// TIA Portal project "e009004v439" (V15.1) (continued)
HMI tags "Tag table_7"
   "Receta Almacén 2\Recetas.REC_MG2.C" : DInt AT %DB51.DBD182, 1 s   // Mot Piece : Côte C
   "Receta Almacén 2\CA_KM01_2" : Bool AT %M19.4, 1 s   // Intercambiador Almacenes Retroceso (Alm2)
   "Receta Almacén 2\OFFSET.REC_MG2.OFFSET_F4" : Int AT %DB52.DBW66, 1 s   // Punto de Formado 4
   "Receta Almacén 2\DB_OP.M2_XCPT" : Bool AT %DB50.DBX382.0, 1 s   // Almacén 2 Entrega Pieza
   "Receta Almacén 2\Detalles" : Bool, internal
   "Receta Almacén 2\DB_OP.M2.MPP" : Bool AT %DB50.DBX420.0, 1 s   // Presencia de Pieza
   "Receta Almacén 2\OFFSET.REC_MG2.OFFSET_F1" : Int AT %DB52.DBW60, 1 s   // Punto de Formado 1
   "Receta Almacén 2\Recetas.REC_MG2.A" : DInt AT %DB51.DBD174, 1 s   // Mot Piece : Côte A
   "Receta Almacén 2\OFFSET.REC_MG2.OFFSET_PL2_1" : Int AT %DB52.DBW72, 1 s   // Plegador 2 Pliego 1
   "Receta Almacén 2\Recetas.REC_MG2.NOM" : String[8] AT %DB51.DBX160.0, 1 s
   "Receta Almacén 2\Recetas.REC_MG2.B" : DInt AT %DB51.DBD178, 1 s   // Mot Piece : Côte B
   "Receta Almacén 2\VerHeladera" : Bool, internal
   "Receta Almacén 2\OFFSET.REC_MG2.OFFSET_F2" : Int AT %DB52.DBW62, 1 s   // Punto de Formado 2
   "Receta Almacén 2\Recetas.REC_MG2.D" : DInt AT %DB51.DBD186, 1 s   // Mot Piece : Côte D
   "Receta Almacén 2\OFFSET.REC_MG2.OFFSET_PL2_2" : Int AT %DB52.DBW74, 1 s   // Plegador 2 Pliego 2
   "Receta Almacén 2\26S6" : Bool AT %I3.5, 1 s   // Presencia de Almacén 2 en Puesto de Espera
   "Receta Almacén 2\OFFSET.REC_MG2.OFFSET_PL1_1" : Int AT %DB52.DBW68, 1 s   // Plegador 1 Pliego 1
   "Receta Almacén 2\OFFSET.REC_MG2.OFFSET_F3" : Int AT %DB52.DBW64, 1 s   // Punto de Formado 3
   "Receta Almacén 2\OFFSET.REC_MG2.OFFSET_PL1_2" : Int AT %DB52.DBW70, 1 s   // Plegador 1 Pliego 2

HMI tags "PiezaPerfiladores"
   "Perfiladores\Perfilador.B" : Int AT %DB8.DBW2, 1 s
   "Perfiladores\Perfilador.PresenciaPieza" : Bool AT %DB8.DBX46.0, 1 s
   "Perfiladores\Perfilador.F1" : Int AT %DB8.DBW8, 1 s
   "Perfiladores\Perfilador.F3" : Int AT %DB8.DBW12, 1 s
   "Perfiladores\Perfilador.PL2_1" : Int AT %DB8.DBW20, 1 s
   "Perfiladores\Perfilador.PL1_1" : Int AT %DB8.DBW16, 1 s
   "Perfiladores\Perfilador.C" : Int AT %DB8.DBW4, 1 s
   "Perfiladores\Perfilador.PL1_2" : Int AT %DB8.DBW18, 1 s
   "Perfiladores\Perfilador.F2" : Int AT %DB8.DBW10, 1 s
   "Perfiladores\Perfilador.F4" : Int AT %DB8.DBW14, 1 s
   "Perfiladores\Perfilador.A" : Int AT %DB8.DBW0, 1 s
   "Perfiladores\Perfilador.PL2_2" : Int AT %DB8.DBW22, 1 s
   "Perfiladores\Perfilador.D" : Int AT %DB8.DBW6, 1 s
   "Forz_Transf-3" : Bool AT %M113.2, 1 s
   "Forz_Transf2" : Bool AT %M113.1, 1 s
   "Forz_Transf1" : Bool AT %M113.0, 1 s
   "Perfiladores\Perfilador.Nombre" : String[20] AT %DB8.DBX24.0, 1 s

HMI tags "PiezaCinta"
   "Cinta\Cinta.PresenciaPieza" : Bool AT %DB9.DBX46.0, 1 s
   "Cinta\Cinta.PL2_1" : Int AT %DB9.DBW20, 1 s
   "Cinta\Cinta.C" : Int AT %DB9.DBW4, 1 s
   "Cinta\Cinta.A" : Int AT %DB9.DBW0, 1 s
   "Cinta\Cinta.F4" : Int AT %DB9.DBW14, 1 s
   "Cinta\Cinta.F3" : Int AT %DB9.DBW12, 1 s
   "Cinta\Cinta.PL2_2" : Int AT %DB9.DBW22, 1 s
   "Cinta\Cinta.PL1_1" : Int AT %DB9.DBW16, 1 s
   "Cinta\Cinta.PL1_2" : Int AT %DB9.DBW18, 1 s
   "Cinta\Cinta.F2" : Int AT %DB9.DBW10, 1 s
   "Cinta\Cinta.D" : Int AT %DB9.DBW6, 1 s
   "Cinta\Cinta.B" : Int AT %DB9.DBW2, 1 s
   "Cinta\Cinta.F1" : Int AT %DB9.DBW8, 1 s
   "Cinta\Cinta.Nombre" : String[20] AT %DB9.DBX24.0, 1 s

HMI tags "PiezaAlm2"
   "Almacén 2\PAlmacén.F3" : Int AT %DB5.DBW12, 1 s
   "Almacén 2\PAlmacén.B" : Int AT %DB5.DBW2, 1 s
   "Almacén 2\PAlmacén.PL2_1" : Int AT %DB5.DBW20, 1 s
   "Almacén 2\PAlmacén.PresenciaPieza" : Bool AT %DB5.DBX46.0, 1 s
   "Almacén 2\PAlmacén.F1" : Int AT %DB5.DBW8, 1 s
   "Almacén 2\PAlmacén.PL2_2" : Int AT %DB5.DBW22, 1 s
   "Almacén 2\PAlmacén.A" : Int AT %DB5.DBW0, 1 s
   "Almacén 2\PAlmacén.F2" : Int AT %DB5.DBW10, 1 s
   "Almacén 2\PAlmacén.F4" : Int AT %DB5.DBW14, 1 s
   "Almacén 2\PAlmacén.C" : Int AT %DB5.DBW4, 1 s
   "Almacén 2\PAlmacén.PL1_1" : Int AT %DB5.DBW16, 1 s
   "Almacén 2\PAlmacén.PL1_2" : Int AT %DB5.DBW18, 1 s
   "Almacén 2\PAlmacén.D" : Int AT %DB5.DBW6, 1 s
   "Almacén 2\PAlmacén.Nombre" : String[20] AT %DB5.DBX24.0, 1 s

HMI tags "PiezaAlm1"
   "Almacén 1\PAlmacén.PL2_2" : Int AT %DB4.DBW22, 1 s
   "Almacén 1\PAlmacén.PL2_1" : Int AT %DB4.DBW20, 1 s
   "Almacén 1\PAlmacén.D" : Int AT %DB4.DBW6, 1 s
   "Almacén 1\PAlmacén.A" : Int AT %DB4.DBW0, 1 s
   "Almacén 1\PAlmacén.F4" : Int AT %DB4.DBW14, 1 s
   "Almacén 1\PAlmacén.B" : Int AT %DB4.DBW2, 1 s
   "Almacén 1\PAlmacén.F3" : Int AT %DB4.DBW12, 1 s
   "Almacén 1\PAlmacén.F2" : Int AT %DB4.DBW10, 1 s
   "Almacén 1\PAlmacén.PL1_2" : Int AT %DB4.DBW18, 1 s
   "Almacén 1\PAlmacén.F1" : Int AT %DB4.DBW8, 1 s
   "Almacén 1\PAlmacén.C" : Int AT %DB4.DBW4, 1 s
   "Almacén 1\PAlmacén.PL1_1" : Int AT %DB4.DBW16, 1 s
   "Almacén 1\PAlmacén.Nombre" : String[20] AT %DB4.DBX24.0, 1 s
   "PL_Resoluc_INCDECF" : Int AT %DB19.DBW8, 1 s
   "PL_Resoluc_INCDECPL" : Int AT %DB19.DBW18, 1 s
   "Almacén 1\PAlmacén.PresenciaPieza_1" : Bool AT %DB4.DBX46.1, 1 s

HMI tags "Alarmas"
   "Alarma 1" : Bool AT %DB50.DBX80.0, 1 s
   "Alarma 2" : Bool AT %DB50.DBX80.1, 1 s
   "Alarma 3" : Bool AT %DB50.DBX80.2, 1 s
   "Alarma 4" : Bool AT %DB50.DBX80.3, 1 s
   "Alarma 5" : Bool AT %DB50.DBX80.4, 1 s
   "Alarma 6" : Bool AT %DB50.DBX80.5, 1 s
   "Alarma 7" : Bool AT %DB50.DBX80.6, 1 s
   "Alarma 8" : Bool AT %DB50.DBX80.7, 1 s
   "Alarma 9" : Bool AT %DB50.DBX81.0, 1 s
   "Alarma 10" : Bool AT %DB50.DBX81.1, 1 s
   "Alarma 11" : Bool AT %DB50.DBX81.2, 1 s
   "Alarma 12" : Bool AT %DB50.DBX81.3, 1 s
   "Alarma 13" : Bool AT %DB50.DBX81.4, 1 s
   "Alarma 14" : Bool AT %DB50.DBX81.5, 1 s
   "Alarma 15" : Bool AT %DB50.DBX81.6, 1 s
   "Alarma 16" : Bool AT %DB50.DBX81.7, 1 s
   "Alarma 17" : Bool AT %DB50.DBX82.0, 1 s
   "Alarma 18" : Bool AT %DB50.DBX82.1, 1 s
   "Alarma 19" : Bool AT %DB50.DBX82.2, 1 s
   "Alarma 20" : Bool AT %DB50.DBX82.3, 1 s
   "Alarma 21" : Bool AT %DB50.DBX82.4, 1 s
   "Alarma 22" : Bool AT %DB50.DBX82.5, 1 s
   "Alarma 23" : Bool AT %DB50.DBX82.6, 1 s
   "Alarma 24" : Bool AT %DB50.DBX82.7, 1 s
   "Alarma 25" : Bool AT %DB50.DBX83.0, 1 s
   "Alarma 26" : Bool AT %DB50.DBX83.1, 1 s
   "Alarma 27" : Bool AT %DB50.DBX83.2, 1 s
   "Alarma 28" : Bool AT %DB50.DBX83.3, 1 s
   "Alarma 29" : Bool AT %DB50.DBX83.4, 1 s
   "Alarma 30" : Bool AT %DB50.DBX83.5, 1 s
   "Alarma 31" : Bool AT %DB50.DBX83.6, 1 s
   "Alarma 32" : Bool AT %DB50.DBX83.7, 1 s
   "Alarma 33" : Bool AT %DB50.DBX84.0, 1 s
   "Alarma 34" : Bool AT %DB50.DBX84.1, 1 s
   "Alarma 35" : Bool AT %DB50.DBX84.2, 1 s
   "Alarma 36" : Bool AT %DB50.DBX84.3, 1 s
   "Alarma 37" : Bool AT %DB50.DBX84.4, 1 s
   "Alarma 38" : Bool AT %DB50.DBX84.5, 1 s
   "Alarma 39" : Bool AT %DB50.DBX84.6, 1 s
   "Alarma 40" : Bool AT %DB50.DBX84.7, 1 s
   "Alarma 41" : Bool AT %DB50.DBX85.0, 1 s
   "Alarma 42" : Bool AT %DB50.DBX85.1, 1 s
   "Alarma 43" : Bool AT %DB50.DBX85.2, 1 s
   "Alarma 44" : Bool AT %DB50.DBX85.3, 1 s
   "Alarma 45" : Bool AT %DB50.DBX85.4, 1 s
   "Alarma 46" : Bool AT %DB50.DBX85.5, 1 s
   "Alarma 47" : Bool AT %DB50.DBX85.6, 1 s
   "Alarma 48" : Bool AT %DB50.DBX85.7, 1 s
   "Alarma 49" : Bool AT %DB50.DBX86.0, 1 s
   "Alarma 50" : Bool AT %DB50.DBX86.1, 1 s
   "Alarma 51" : Bool AT %DB50.DBX86.2, 1 s
   "Alarma 52" : Bool AT %DB50.DBX86.3, 1 s
   "Alarma 53" : Bool AT %DB50.DBX86.4, 1 s
   "Alarma 54" : Bool AT %DB50.DBX86.5, 1 s
   "Alarma 55" : Bool AT %DB50.DBX86.6, 1 s
   "Alarma 56" : Bool AT %DB50.DBX86.7, 1 s
   "Alarma 57" : Bool AT %DB50.DBX87.0, 1 s
   "Alarma 58" : Bool AT %DB50.DBX87.1, 1 s
   "Alarma 59" : Bool AT %DB50.DBX87.2, 1 s
   "Alarma 60" : Bool AT %DB50.DBX87.3, 1 s
   "Alarma 61" : Bool AT %DB50.DBX87.4, 1 s
   "Alarma 62" : Bool AT %DB50.DBX87.5, 1 s
   "Alarma 63" : Bool AT %DB50.DBX87.6, 1 s
   "Alarma 64" : Bool AT %DB50.DBX87.7, 1 s
   "Alarma 65" : Bool AT %DB50.DBX88.0, 1 s
   "Alarma 66" : Bool AT %DB50.DBX88.1, 1 s
   "Alarma 67" : Bool AT %DB50.DBX88.2, 1 s
   "Alarma 68" : Bool AT %DB50.DBX88.3, 1 s
   "Alarma 69" : Bool AT %DB50.DBX88.4, 1 s
   "Alarma 70" : Bool AT %DB50.DBX88.5, 1 s
   "Alarma 71" : Bool AT %DB50.DBX88.6, 1 s
   "Alarma 72" : Bool AT %DB50.DBX88.7, 1 s
   "Alarma 73" : Bool AT %DB50.DBX89.0, 1 s
   "Alarma 74" : Bool AT %DB50.DBX89.1, 1 s
   "Alarma 75" : Bool AT %DB50.DBX89.2, 1 s
   "Alarma 76" : Bool AT %DB50.DBX89.3, 1 s
   "Alarma 77" : Bool AT %DB50.DBX89.4, 1 s
   "Alarma 78" : Bool AT %DB50.DBX89.5, 1 s
   "Alarma 79" : Bool AT %DB50.DBX89.6, 1 s
   "Alarma 80" : Bool AT %DB50.DBX89.7, 1 s
   "Alarma 81" : Bool AT %DB50.DBX90.0, 1 s
   "Alarma 82" : Bool AT %DB50.DBX90.1, 1 s
   "Alarma 83" : Bool AT %DB50.DBX90.2, 1 s
   "Alarma 84" : Bool AT %DB50.DBX90.3, 1 s
   "Alarma 85" : Bool AT %DB50.DBX90.4, 1 s
   "Alarma 86" : Bool AT %DB50.DBX90.5, 1 s
   "Alarma 87" : Bool AT %DB50.DBX90.6, 1 s
   "Alarma 88" : Bool AT %DB50.DBX90.7, 1 s
   "Alarma 89" : Bool AT %DB50.DBX91.0, 1 s
   "Alarma 90" : Bool AT %DB50.DBX91.1, 1 s
   "Alarma 91" : Bool AT %DB50.DBX91.2, 1 s
   "Alarma 92" : Bool AT %DB50.DBX91.3, 1 s
   "Alarma 93" : Bool AT %DB50.DBX91.4, 1 s
   "Alarma 94" : Bool AT %DB50.DBX91.5, 1 s
   "Alarma 95" : Bool AT %DB50.DBX91.6, 1 s
   "Alarma 96" : Bool AT %DB50.DBX91.7, 1 s
   "Alarma 97" : Bool AT %DB50.DBX92.0, 1 s
   "Alarma 98" : Bool AT %DB50.DBX92.1, 1 s
   "Alarma 99" : Bool AT %DB50.DBX92.2, 1 s
   "Alarma 100" : Bool AT %DB50.DBX92.3, 1 s
   "Alarma 101" : Bool AT %DB50.DBX92.4, 1 s
   "Alarma 102" : Bool AT %DB50.DBX92.5, 1 s
   "Alarma 103" : Bool AT %DB50.DBX92.6, 1 s
   "Alarma 104" : Bool AT %DB50.DBX92.7, 1 s
   "Alarma 105" : Bool AT %DB50.DBX93.0, 1 s
   "Alarma 106" : Bool AT %DB50.DBX93.1, 1 s
   "Alarma 107" : Bool AT %DB50.DBX93.2, 1 s
   "Alarma 108" : Bool AT %DB50.DBX93.3, 1 s
   "Alarma 109" : Bool AT %DB50.DBX93.4, 1 s
   "Alarma 110" : Bool AT %DB50.DBX93.5, 1 s
   "Alarma 111" : Bool AT %DB50.DBX93.6, 1 s
   "Alarma 112" : Bool AT %DB50.DBX93.7, 1 s
   "Alarma 113" : Bool AT %DB50.DBX94.0, 1 s
   "Alarma 114" : Bool AT %DB50.DBX94.1, 1 s
   "Alarma 115" : Bool AT %DB50.DBX94.2, 1 s
   "Alarma 116" : Bool AT %DB50.DBX94.3, 1 s
   "Alarma 117" : Bool AT %DB50.DBX94.4, 1 s
   "Alarma 118" : Bool AT %DB50.DBX94.5, 1 s
   "Alarma 119" : Bool AT %DB50.DBX94.6, 1 s
   "Alarma 120" : Bool AT %DB50.DBX94.7, 1 s
   "Alarma 121" : Bool AT %DB50.DBX95.0, 1 s
   "PL1_Pos00" : Bool AT %DB50.DBX393.0, 1 s

HMI tags "Atasco Perfilador"
   "Sensor 1" : Bool AT %I14.4, 100 ms
   "Sensor 2" : Bool AT %I14.5, 100 ms
   "Sensor 3" : Bool AT %I14.6, 100 ms
   "Sensor 4" : Bool AT %I14.7, 100 ms
   "Sensor 5" : Bool AT %I18.3, 100 ms
   "Sensor 6" : Bool AT %I16.0, 100 ms
   "Sensor 7" : Bool AT %I16.1, 100 ms
   "Sensor 8" : Bool AT %I16.2, 100 ms
   "Sensor 9" : Bool AT %I16.3, 100 ms
   "Sensor 10" : Bool AT %I16.4, 100 ms
   "Sensor 11" : Bool AT %I16.5, 100 ms
   "Sensor 12" : Bool AT %I16.6, 100 ms
   "Sensor 13" : Bool AT %I16.7, 100 ms
   "Sensor 14" : Bool AT %I17.0, 100 ms
   "Sensor 15" : Bool AT %I17.1, 100 ms
   "Sensor 16" : Bool AT %I17.2, 100 ms
   "Sensor 17" : Bool AT %I17.3, 100 ms
   "Sensor 18" : Bool AT %I17.4, 100 ms
   "Sensor 19" : Bool AT %I17.5, 100 ms
   "Sensor 20" : Bool, internal
   "Sensor 21" : Bool AT %I17.6, 100 ms
   "Sensor 22" : Bool AT %I18.0, 100 ms
   "Sensor 23" : Bool AT %I18.1, 100 ms
   "Sensor 24" : Bool AT %I18.2, 100 ms
   "36S10" : Bool AT %I15.0, 1 s

HMI tags "PiezaDescargador"
   "Descargador-A" : Int AT %DB12.DBW0, 1 s
   "Descargador-B" : Int AT %DB12.DBW2, 1 s
   "Descargador-C" : Int AT %DB12.DBW4, 1 s
   "Descargador-D" : Int AT %DB12.DBW6, 1 s
   "Descargador-F1" : Int AT %DB12.DBW8, 1 s
   "Descargador-F2" : Int AT %DB12.DBW10, 1 s
   "Descargador-F3" : Int AT %DB12.DBW12, 1 s
   "Descargador-F4" : Int AT %DB12.DBW14, 1 s
   "Descargador-PL1_1" : Int AT %DB12.DBW16, 1 s
   "Descargador-PL1_2" : Int AT %DB12.DBW18, 1 s
   "Descargador-PL2_1" : Int AT %DB12.DBW20, 1 s
   "Descargador-PL2_2" : Int AT %DB12.DBW22, 1 s
   "Descargador-Nombre" : String[20] AT %DB12.DBX24.0, 1 s
   "Descargador-PiezaPresente" : Bool AT %DB12.DBX46.0, 1 s
   "Descargador-Almacen" : Bool AT %DB12.DBX46.1, 1 s
   "Descargador-PL2_3" : Int AT %DB12.DBW24, 1 s

HMI tags "ProcesoPlegadores"
   "PL_Estados" : Int AT %MW150, 1 s
   "PL_Concatenadoras" : Int AT %MW152, 1 s
   "PL_S_0" : Bool AT %M150.0, 1 s
   "PL_S_1" : Bool AT %M150.1, 1 s
   "PL_S_2" : Bool AT %M150.2, 1 s
   "PL_S_3" : Bool AT %M150.3, 1 s
   "PL_S_4" : Bool AT %M150.4, 1 s
   "PL_S_5" : Bool AT %M150.5, 1 s
   "PL_S_6" : Bool AT %M150.6, 1 s
   "PL_S_7" : Bool AT %M150.7, 1 s
   "PL_S_8" : Bool AT %M151.0, 1 s
   "PL_S_9" : Bool AT %M151.1, 1 s
   "PL_S_10" : Bool AT %M151.2, 1 s
   "PL_S_11" : Bool AT %M151.3, 1 s
   "PL_S_12" : Bool AT %M151.4, 1 s
   "PL_S_13" : Bool AT %M151.5, 1 s
   "PL_S_14" : Bool AT %M151.6, 1 s
   "PL_S_15" : Bool AT %M151.7, 1 s
   "STOP_RUN" : Bool AT %M101.3, 1 s
   "PL_Continuar" : Bool AT %M101.4, 1 s
   "PL_Reset" : Bool AT %M101.5, 1 s
   "PL_en_Ciclo" : Bool AT %M10.3, 1 s
   "PL_Prioritarias" : Int AT %MW154, 1 s
   "PL_P_0" : Bool AT %M154.0, 1 s
   "PL_P_1" : Bool AT %M154.1, 1 s
   "PL_P_2" : Bool AT %M154.2, 1 s
   "PL_P_3" : Bool AT %M154.3, 1 s
   "PL_P_4" : Bool AT %M154.4, 1 s
   "PL_P_5" : Bool AT %M154.5, 1 s
   "PL_P_6" : Bool AT %M154.6, 1 s
   "PL_P_7" : Bool AT %M154.7, 1 s
   "PL_P_8" : Bool AT %M155.0, 1 s
   "PL_P_9" : Bool AT %M155.1, 1 s
   "PL_P_10" : Bool AT %M155.2, 1 s
   "PL_P_11" : Bool AT %M155.3, 1 s
   "PL_P_12" : Bool AT %M155.4, 1 s
   "PL_P_13" : Bool AT %M155.5, 1 s
   "PL_P_14" : Bool AT %M155.6, 1 s
   "PL_P_15" : Bool AT %M155.7, 1 s
   "PL_Req_Pos_Recep" : Bool AT %M100.0, 1 s
   "PL_Req_Pos_Pleg1" : Bool AT %M100.1, 1 s
   "PL_Req_Pos_Pleg2" : Bool AT %M100.3, 1 s
   "PL_Req_Pos_Entrega" : Bool AT %M100.4, 1 s
   "PL_Req_Pos_Espera" : Bool AT %M100.5, 1 s
   "PL_En_Pos_Espera" : Bool AT %M180.0, 1 s
   "PL_En_Pos_Recepción" : Bool AT %M180.1, 1 s
   "PL_En_Pos_Pleg1" : Bool AT %M180.3, 1 s
   "PL_En_Pos_Pleg2" : Bool AT %M180.4, 1 s
   "PL_En_Pos_Entrega" : Bool AT %M180.5, 1 s
   "PL_MovimientoSeguro" : Bool AT %M181.1, 1 s
   "PL_Prensas_No" : Bool AT %M165.5, 1 s
   "PL_Fijaciones_No" : Bool AT %M165.7, 1 s
   "PL_Alineado_No" : Bool AT %M165.1, 1 s
   "PL_Cepillos_No" : Bool AT %M165.3, 1 s
   "PL_Plegado_No" : Bool AT %M170.3, 1 s
   "PL_Simu1_PrensaNo" : Bool AT %M55.0, 1 s
   "PL_Simu2_AliNo" : Bool AT %M55.1, 1 s
   "PL_Simu3_CepNo" : Bool AT %M55.2, 1 s
   "PL_Simu4_FijaNo" : Bool AT %M55.3, 1 s
   "PL_Simu5_PlegNo" : Bool AT %M55.4, 1 s
   "PL_Alineado_SI" : Bool AT %M165.0, 1 s
   "PL_Cepillos_SI" : Bool AT %M165.2, 1 s
   "PL_Prensas_SI" : Bool AT %M165.4, 1 s
   "PL_Fijaciones_SI" : Bool AT %M165.6, 1 s
   "PL_Plegador1_ON" : Bool AT %M166.0, 1 s
   "PL_Plegador2_ON" : Bool AT %M166.2, 1 s
   "PL_Tenaza_Arriba" : Bool AT %M170.5, 1 s
   "PL_Tenaza_Abajo" : Bool AT %M170.6, 1 s
   "PL_Tenaza_Abierta" : Bool AT %M170.7, 1 s
   "PL_Tenaza_Cerrada" : Bool AT %M171.0, 1 s
   "PL_Tenaza_Adelante" : Bool AT %M171.1, 1 s
   "PL_Tenaza_Atrás" : Bool AT %M171.2, 1 s
   "PL_Desc_Adelante" : Bool AT %M171.3, 1 s
   "PL_Desc_Atrás" : Bool AT %M171.4, 1 s
   "PL_Dec_F_A1" : Int AT %DB19.DBW2, 1 s
   "PL_Inc_F_A1" : Int AT %DB19.DBW0, 1 s
   "PL_Dec_F_A2" : Int AT %DB19.DBW6, 1 s
   "PL_Inc_F_A2" : Int AT %DB19.DBW4, 1 s
   "PL_Inc_PL_A1" : Int AT %DB1.DBW10, 1 s
   "PL_Dec_PL_A1" : Int AT %DB19.DBW12, 1 s
   "PL_Inc_PL_A2" : Int AT %DB19.DBW14, 1 s
   "PL_Dec_PL_A2" : Int AT %DB19.DBW16, 1 s

HMI tags "ReferenciasServos"
   "PosiciónEspera_PL1" : DInt AT %DB55.DBD8, 1 s
   "PosiciónRecepción_PL1" : DInt AT %DB55.DBD12, 1 s
   "PosiciónPlegado1_PL1" : DInt AT %DB55.DBD16, 1 s
   "PosiciónPlegado2_PL1" : DInt AT %DB55.DBD20, 1 s
   "PosiciónEntrega_PL1" : DInt AT %DB55.DBD24, 1 s
   "PosiciónEspera_PL2" : DInt AT %DB54.DBD8, 1 s
   "PosiciónRecepción_PL2" : DInt AT %DB54.DBD12, 1 s
   "PosiciónPlegado1_PL2" : DInt AT %DB54.DBD16, 1 s
   "PosiciónPlegado2_PL2" : DInt AT %DB54.DBD20, 1 s
   "PosiciónEntrega_PL2" : DInt AT %DB54.DBD24, 1 s
   "PosiciónMínima_PL" : DInt AT %DB16.DBD24, 1 s
   "PosiciónMáxima_PL" : DInt AT %DB16.DBD20, 1 s
   "PosiciónActual_PL1" : DInt AT %DB50.DBD200, 1 s
   "PosiciónActual_PL2" : DInt AT %DB50.DBD250, 1 s
   "PosiciónRecepción_PL2(Ant)" : DInt AT %DB58.DBD12, 1 s
   "PosiciónPlegado1_PL2(Ant)" : DInt AT %DB58.DBD16, 1 s
   "PosiciónPlegado2_PL2(Ant)" : DInt AT %DB58.DBD20, 1 s
   "PosiciónEntrega_PL2(Ant)" : DInt AT %DB58.DBD24, 1 s
   "PosiciónEspera_PL2(Ant)" : DInt AT %DB58.DBD8, 1 s
   "PosiciónRecepción_PL1(Ant)" : DInt AT %DB57.DBD12, 1 s
   "PosiciónPlegado1_PL1(Ant)" : DInt AT %DB57.DBD16, 1 s
   "PosiciónPlegado2_PL1(Ant)" : DInt AT %DB57.DBD20, 1 s
   "PosiciónEntrega_PL1(Ant)" : DInt AT %DB57.DBD24, 1 s
   "PosiciónEspera_PL1(Ant)" : DInt AT %DB57.DBD8, 1 s

HMI tags "ProcesoPinza"
   "F_Concatenadoras" : Int AT %MW206, 1 s
   "F_C_0" : Bool AT %M206.0, 1 s
   "F_C_1" : Bool AT %M206.1, 1 s
   "F_C_2" : Bool AT %M206.2, 1 s
   "F_C_3" : Bool AT %M206.3, 1 s
   "F_C_4" : Bool AT %M206.4, 1 s
   "F_C_5" : Bool AT %M206.5, 1 s
   "F_C_6" : Bool AT %M206.6, 1 s
   "F_C_7" : Bool AT %M206.7, 1 s
   "F_C_8" : Bool AT %M207.0, 1 s
   "F_C_9" : Bool AT %M207.1, 1 s
   "F_C_10" : Bool AT %M207.2, 1 s
   "F_C_11" : Bool AT %M207.3, 1 s
   "F_C_12" : Bool AT %M207.4, 1 s
   "F_C_13" : Bool AT %M207.5, 1 s
   "F_C_14" : Bool AT %M207.6, 1 s
   "F_C_15" : Bool AT %M207.7, 1 s
   "F_P_0" : Bool AT %M208.0, 1 s
   "F_P_1" : Bool AT %M208.1, 1 s
   "F_P_2" : Bool AT %M208.2, 1 s
   "F_P_3" : Bool AT %M208.3, 1 s
   "F_P_4" : Bool AT %M208.4, 1 s
   "F_P_5" : Bool AT %M208.5, 1 s
   "F_P_6" : Bool AT %M208.6, 1 s
   "F_P_7" : Bool AT %M208.7, 1 s
   "F_P_8" : Bool AT %M209.0, 1 s
   "F_P_9" : Bool AT %M209.1, 1 s
   "F_P_10" : Bool AT %M209.2, 1 s
   "F_P_11" : Bool AT %M209.3, 1 s
   "F_P_12" : Bool AT %M209.4, 1 s
   "F_P_13" : Bool AT %M209.5, 1 s
   "F_P_14" : Bool AT %M209.6, 1 s
   "F_P_15" : Bool AT %M209.7, 1 s
   "F_S_0" : Bool AT %M204.0, 1 s
   "F_S_1" : Bool AT %M204.1, 1 s
   "F_S_2" : Bool AT %M204.2, 1 s
   "F_S_3" : Bool AT %M204.3, 1 s
   "F_S_4" : Bool AT %M204.4, 1 s
   "F_S_5" : Bool AT %M204.5, 1 s
   "F_S_6" : Bool AT %M204.6, 1 s
   "F_S_7" : Bool AT %M204.7, 1 s
   "F_S_8" : Bool AT %M205.0, 1 s
   "F_S_9" : Bool AT %M205.1, 1 s
   "F_S_10" : Bool AT %M205.2, 1 s
   "F_S_11" : Bool AT %M205.3, 1 s
   "F_S_12" : Bool AT %M205.4, 1 s
   "F_S_13" : Bool AT %M205.5, 1 s
   "F_S_14" : Bool AT %M205.6, 1 s
   "F_S_15" : Bool AT %M205.7, 1 s
   "F_Estados" : Int AT %MW204, 1 s
   "F_H1_No" : Bool AT %M210.7, 1 s
   "F_H2_No" : Bool AT %M211.1, 1 s
   "F_MovimientoSeguro" : Bool AT %M181.2, 1 s
   "F_Tenaza_No" : Bool AT %M171.2, 1 s
   "F_Descargador_No" : Bool AT %I8.2, 1 s
   "F_SimuH1_No" : Bool AT %M58.0, 1 s
   "F_SimuH2_No" : Bool AT %M58.1, 1 s
   "F_SimuTenaza_No" : Bool AT %M58.2, 1 s
   "F_Req_Pos_Espera" : Bool AT %M104.5, 1 s
   "F_Req_Pos_E1H1" : Bool AT %M104.0, 1 s
   "F_Req_Pos_E1H2" : Bool AT %M104.1, 1 s
   "F_Req_Pos_E2H1" : Bool AT %M104.2, 1 s
   "F_Req_Pos_E2H2" : Bool AT %M104.3, 1 s
   "F_Req_Pos_Entrega" : Bool AT %M104.4, 1 s
   "F_En_Pos_Espera" : Bool AT %DB50.DBX392.0, 1 s
   "F_En_Pos_E1H1" : Bool AT %DB50.DBX392.1, 1 s
   "F_En_Pos_E1H2" : Bool AT %DB50.DBX392.2, 1 s
   "F_En_Pos_E2H1" : Bool AT %DB50.DBX392.3, 1 s
   "F_En_Pos_E2H2" : Bool AT %DB50.DBX392.4, 1 s
   "F_En_Pos_Entrega" : Bool AT %DB50.DBX392.5, 1 s

HMI tags "ReferenciasServo"
   "PosiciónEspera_F" : DInt AT %DB13.DBD0, 1 s
   "PosiciónE1H1_F" : DInt AT %DB13.DBD4, 1 s
   "PosiciónE1H2_F" : DInt AT %DB13.DBD8, 1 s
   "PosiciónE2H1_F" : DInt AT %DB13.DBD12, 1 s
   "PosiciónE2H2_F" : DInt AT %DB13.DBD16, 1 s
   "PosiciónEntrega_F" : DInt AT %DB13.DBD20, 1 s
   "PosiciónMáxima_F" : DInt AT %DB16.DBD16, 1 s
   "PosiciónActual_F" : DInt AT %DB50.DBD300, 1 s
   "F_Referencia_Menor_Descargador" : Bool AT %M57.0, 1 s
   "Distancia_entre_Herramientas_F" : DInt AT %DB16.DBD0, 1 s
   "Distancia_entre_Herramienta1_y_Pos0_F" : DInt AT %DB16.DBD4, 1 s
   "Distancia_entre_Pos0_y_Tenaza_F" : DInt AT %DB16.DBD8, 1 s
   "Distancia_entre_Pos0_y_Descargador_F" : DInt AT %DB16.DBD12, 1 s
   "PosiciónE1H1_F(Ant)" : DInt AT %DB18.DBD4, 1 s
   "PosiciónE1H2_F(Ant)" : DInt AT %DB18.DBD8, 1 s
   "PosiciónE2H1_F(Ant)" : DInt AT %DB18.DBD12, 1 s
   "PosiciónE2H2_F(Ant)" : DInt AT %DB18.DBD16, 1 s
   "PosiciónEntrega_F(Ant)" : DInt AT %DB18.DBD20, 1 s
   "PosiciónEspera_F(Ant)" : DInt AT %DB18.DBD0, 1 s
   "Distancia_entre_Pleg_Alin_PL" : DInt AT %DB16.DBD28, 1 s

HMI tags "Registro de Pos"
   "Pos_Recepcion" : DInt AT %DB18.DBD0, 1 s   // "Posiciones_Pinza_Ant".Pos_Recepcion
   "Pos_E1H1" : DInt AT %DB18.DBD4, 1 s   // "Posiciones_Pinza_Ant".Pos_E1H1
   "Pos_E1H2" : DInt AT %DB18.DBD8, 1 s   // "Posiciones_Pinza_Ant".Pos_E1H2
   "Pos_E2H1" : DInt AT %DB18.DBD12, 1 s   // "Posiciones_Pinza_Ant".Pos_E2H1
   "Pos_E2H2" : DInt AT %DB18.DBD16, 1 s   // "Posiciones_Pinza_Ant".Pos_E2H2
   "Pos_Entrega" : DInt AT %DB18.DBD20, 1 s   // "Posiciones_Pinza_Ant".Pos_Entrega
   "Pos_Recepcion(1)" : DInt AT %DB23.DBD0, 1 s   // "Posiciones_Pinza_Ant2".Pos_Recepcion
   "Pos_E1H1(1)" : DInt AT %DB23.DBD4, 1 s   // "Posiciones_Pinza_Ant2".Pos_E1H1
   "Pos_E1H2(1)" : DInt AT %DB23.DBD8, 1 s   // "Posiciones_Pinza_Ant2".Pos_E1H2
   "Pos_E2H1(1)" : DInt AT %DB23.DBD12, 1 s   // "Posiciones_Pinza_Ant2".Pos_E2H1
   "Pos_E2H2(1)" : DInt AT %DB23.DBD16, 1 s   // "Posiciones_Pinza_Ant2".Pos_E2H2
   "Pos_Entrega(1)" : DInt AT %DB23.DBD20, 1 s   // "Posiciones_Pinza_Ant2".Pos_Entrega
   "Pos_Recepcion(2)" : DInt AT %DB24.DBD0, 1 s   // "Posiciones_Pinza_Ant3".Pos_Recepcion
   "Pos_E1H1(2)" : DInt AT %DB24.DBD4, 1 s   // "Posiciones_Pinza_Ant3".Pos_E1H1
   "Pos_E1H2(2)" : DInt AT %DB24.DBD8, 1 s   // "Posiciones_Pinza_Ant3".Pos_E1H2
   "Pos_E2H1(2)" : DInt AT %DB24.DBD12, 1 s   // "Posiciones_Pinza_Ant3".Pos_E2H1
   "Pos_E2H2(2)" : DInt AT %DB24.DBD16, 1 s   // "Posiciones_Pinza_Ant3".Pos_E2H2
   "Pos_Entrega(2)" : DInt AT %DB24.DBD20, 1 s   // "Posiciones_Pinza_Ant3".Pos_Entrega
   "Pos_Recepcion(3)" : DInt AT %DB26.DBD0, 1 s   // "PosReal_Pinza_Ant".Pos_Recepcion
   "Pos_E1H1(3)" : DInt AT %DB26.DBD4, 1 s   // "PosReal_Pinza_Ant".Pos_E1H1
   "Pos_E1H2(3)" : DInt AT %DB26.DBD8, 1 s   // "PosReal_Pinza_Ant".Pos_E1H2
   "Pos_E2H1(3)" : DInt AT %DB26.DBD12, 1 s   // "PosReal_Pinza_Ant".Pos_E2H1
   "Pos_E2H2(3)" : DInt AT %DB26.DBD16, 1 s   // "PosReal_Pinza_Ant".Pos_E2H2
   "Pos_Entrega(3)" : DInt AT %DB26.DBD20, 1 s   // "PosReal_Pinza_Ant".Pos_Entrega
   "Pos_Recepcion(4)" : DInt AT %DB27.DBD0, 1 s   // "PosReal_Pinza_Ant2".Pos_Recepcion
   "Pos_E1H1(4)" : DInt AT %DB27.DBD4, 1 s   // "PosReal_Pinza_Ant2".Pos_E1H1
   "Pos_E1H2(4)" : DInt AT %DB27.DBD8, 1 s   // "PosReal_Pinza_Ant2".Pos_E1H2
   "Pos_E2H1(4)" : DInt AT %DB27.DBD12, 1 s   // "PosReal_Pinza_Ant2".Pos_E2H1
   "Pos_E2H2(4)" : DInt AT %DB27.DBD16, 1 s   // "PosReal_Pinza_Ant2".Pos_E2H2
   "Pos_Entrega(4)" : DInt AT %DB27.DBD20, 1 s   // "PosReal_Pinza_Ant2".Pos_Entrega
   "Pos_Recepcion(5)" : DInt AT %DB28.DBD0, 1 s   // "PosReal_Pinza_Ant3".Pos_Recepcion
   "Pos_E1H1(5)" : DInt AT %DB28.DBD4, 1 s   // "PosReal_Pinza_Ant3".Pos_E1H1
   "Pos_E1H2(5)" : DInt AT %DB28.DBD8, 1 s   // "PosReal_Pinza_Ant3".Pos_E1H2
   "Pos_E2H1(5)" : DInt AT %DB28.DBD12, 1 s   // "PosReal_Pinza_Ant3".Pos_E2H1
   "Pos_E2H2(5)" : DInt AT %DB28.DBD16, 1 s   // "PosReal_Pinza_Ant3".Pos_E2H2
   "Pos_Entrega(5)" : DInt AT %DB28.DBD20, 1 s   // "PosReal_Pinza_Ant3".Pos_Entrega
   "Pos_Recepcion(6)" : DInt AT %DB29.DBD0, 1 s   // "Error_Pinza_Ant".Pos_Recepcion
   "Pos_E1H1(6)" : DInt AT %DB29.DBD4, 1 s   // "Error_Pinza_Ant".Pos_E1H1
   "Pos_E1H2(6)" : DInt AT %DB29.DBD8, 1 s   // "Error_Pinza_Ant".Pos_E1H2
   "Pos_E2H1(6)" : DInt AT %DB29.DBD12, 1 s   // "Error_Pinza_Ant".Pos_E2H1
   "Pos_E2H2(6)" : DInt AT %DB29.DBD16, 1 s   // "Error_Pinza_Ant".Pos_E2H2
   "Pos_Entrega(6)" : DInt AT %DB29.DBD20, 1 s   // "Error_Pinza_Ant".Pos_Entrega

discrete alarms
   83: 'Falla al abrir pinza posicionadora: Comprobar Sensores 29S4 y 29S5 + Electroválvula 43Y7 / FORMAGE : DEF MOUVEMENT OUVERTURE PINCE 43Y7 : vérifier 29S4 29S5', class Fallos Pinza, trigger "DB_OP.DEF06" bit 10
   41: 'Falla retroceso de pinza en Plegadora: Comprobar Sensores 30S1 y 30S2 + Electroválvula 44Y2 / PLIEUSE : DEF MOUVEMENT RECUL PINCE 44Y2 : vérifier 30S1 et 30S2', class Fallos Plegadora, trigger "DB_OP.DEF03" bit 0
   35: 'Falla al abrir pinza en Plegadora: Comprobar Sensores 30S5 y 30S6 + Electroválvula 44Y5 / PLIEUSE : DEF MOUVEMENT OUVERTURE PINCE 44Y5 : vérifier 30S5 et 30S6', class Fallos Plegadora, trigger "DB_OP.DEF03" bit 10
   112: 'Reserva', class Reserva, trigger "DB_OP.DEF07" bit 7
   85: 'Falla al retroceder ajuste de formado: Comprobar Contactor KM09.2 + Encóder correspondiente / FORMAGE : DEF MOUVEMENT RECUL MOP KM09_2 : vérifier codeur 2', class Fallos Formado, trigger "DB_OP.DEF06" bit 12
   62: 'Falla en Plegador 2 al intentar desactivar orden de plegado: Comprobar Sensores 35S3 y 35S4 + Relé 47K4 / PLIEUSE 1 : DEF MOUVEMENT RECUL PLIAGE 45K6 : vérifier 31S7 et 31S8', class Fallos Plegadora, trigger "DB_OP.DEF04" bit 5
   100: 'Falla al retroceder matriz de herramienta 2 en Formador: Comprobar Sensores 28S3 y 28S4 + Relé43K2 / FORMAGE : DEF MOUVEMENT RECUL MATRICE OUTIL 2 43K2 : vérifier 28S3 28S4', class Fallos Formado, trigger "DB_OP.DEF07" bit 11
   74: 'Se intentó bajar la araña a traves de la electroválvula 41Y1, pero no se recibe la confirmación adecuada del sensor 26S1. / Falla al bajar Araña: Comprobar Sensor 26S1, y Electroválvula 41Y1 / PREHENSEUR : DEF MOUVEMENT DESCENTE 41Y1 : vérifier', class Fallos Araña, trigger "DB_OP.DEF05" bit 1
   28: 'Falla Temperatura Grupo Hidráulico: Comprobar Termostato 23S8 / DEFAUT TEMPERATURE GROUPE HYDRAULIQUE', class Fallos Generales, trigger "DB_OP.DEF02" bit 3
   91: 'Falla al avanzar martillo de herramienta 2 en Formador: Comprobar Sensores 28S1 y 28S2 + Relé 42K7 / FORMAGE : DEF MOUVEMENT AVANCE MARTEAU OUTIL 2 42K7 : vérifier 28S1 28S2', class Fallos Formado, trigger "DB_OP.DEF06" bit 2
   103: 'Falla al retroceder intercambiador de Almacenes: Comprobar Sensores 26S6 y 26S7 + Contactor KM01.2 / CHARGEMENT : DEF MOUVEMENT RECUL MAGASIN : vérifier 26S6 26S7', class Fallos Almacenes, trigger "DB_OP.DEF07" bit 14
   61: 'Falla en Plegador 2 al intentar desactivar fijación: Comprobar Sensores 35S1 y 35S2 + Relé 47K2', class Fallos Plegadora, trigger "DB_OP.DEF04" bit 4
   49: 'Falla en Plegador 1 al intentar activar fijación: Comprobar Sensores 31S5 y 31S6 + Relé 45K3 / PLIEUSE 1 : DEF MOUVEMENT AVANCE BRIDAGE 45K3 : vérifier 31S5 et 31S6', class Fallos Plegadora, trigger "DB_OP.DEF04" bit 8
   33: 'Falla avance de pinza en Plegadora: Comprobar Sensores 30S1 y 30S2 + Electroválvula 44Y1 / PLIEUSE : DEF MOUVEMENT AVANCE PINCE 44Y1 : vérifier 30S1 et 30S2', class Fallos Plegadora, trigger "DB_OP.DEF03" bit 8
   90: 'Falla al avanzar matriz de herramienta 1 en Formador: Comprobar Sensores 27S7 y 27S8 + Relé 42K5 / FORMAGE : DEF MOUVEMENT AVANCE MATRICE OUTIL 1 42K5 : vérifier 27S7 27S8', class Fallos Formado, trigger "DB_OP.DEF06" bit 1
   113: 'Reserva', class Reserva, trigger "DB_OP.DEF08" bit 8
   82: 'Falla al subir Bloqueador de Avance en etapa formador: Comprobar Sensores 29S1 y 29S2 + Electroválula 43Y6 / FORMAGE : DEF MOUVEMENT MONTEE BUTEE 43Y6 : vérifier 29S1 29S2', class Fallos Formado, trigger "DB_OP.DEF06" bit 9
   3: 'Falla Alimentación Motor Intercambio de Almacenes: Comprobar estado de Guardamotor QM01 / Moteur OK Axe Magasin Tôle', class Fallos Almacenes, trigger "DB_OP.DEF01" bit 10
   2: 'Falla Almacenes Deshabilitados / Réchauffeur Tôle OK (option)', class Fallos Almacenes, trigger "DB_OP.DEF01" bit 9
   14: 'Falla térmica en motor ajuste de ancho en etapa de formado: Comprobar estado de Guardamotor QM09 / DF_QM09 : FORMAGE : Moteur OK Axe', class Fallos Generales, trigger "DB_OP.DEF01" bit 5
   117: 'Reserva', class Reserva, trigger "DB_OP.DEF08" bit 12
   29: 'Falla Seguridad Barrera en Descargador: Comprobar estado de Sensor 31S4 / DEFAUT BARRIERE', class Fallos Descargador, trigger "DB_OP.DEF02" bit 4
   55: 'Falla en Plegador 2 al intentar bajar prensa: Comprobar Sensores 35S5 y 35S6 + Relé 45K5 / PLIEUSE 1 : DEF MOUVEMENT AVANCE V1 45K7 : vérifier 32S1 et 32S2', class Fallos Plegadora, trigger "DB_OP.DEF04" bit 14
   30: 'Falla Cubierta de Perfilador: Comprobar Sensor 34S1 / DEFAUT CARTER PROFILEUSE', class Fallos Perfiladores, trigger "DB_OP.DEF02" bit 5
   121: 'Inconsistencia de Presencia de pieza en en Descargador: Comprobar Sensor 31S1 / DECHARGEMENT : defaut presence piece', class Fallos Descargador, trigger "DB_OP.DEF08" bit 0
   116: 'Inconsistencia de Presencia de pieza en Transporte de Rolos: Comprobar Sensor 26S8 / Convoyeur 1 : defaut presence piece', class Fallos Rolos, trigger "DB_OP.DEF08" bit 11
   66: 'Se intentó subir la araña a traves de la electroválvula 40Y7, pero no se recibe la confirmación adecuada del sensor 25S4. / Falla al subir Araña: Comprobar sensor 25S4 + Electroválvula 40Y7 / PREHENSEUR : DEF MOUVEMENT MONTEE 40Y7 : vérifier 25S4', class Fallos Araña, trigger "DB_OP.DEF05" bit 9
   51: 'Falla en Plegador 1 al intentar bajar prensa: Comprobar Sensores 32S1 y 32S2 + Relé 45K7 / PLIEUSE 1 : DEF MOUVEMENT AVANCE V1 45K7 : vérifier 32S1 et 32S2', class Fallos Plegadora, trigger "DB_OP.DEF04" bit 10
   70: 'Reserva', class Reserva, trigger "DB_OP.DEF05" bit 13
   64: 'Falla en Plegador 2 al intentar subir primera extensión de prensa: Comprobar Sensores 35S7 y 35S8 + Relé 46K8 / PLIEUSE 2 : DEF MOUVEMENT AVANCE V2 47K7 : vérifier 35S7 et 35S8', class Fallos Plegadora, trigger "DB_OP.DEF04" bit 7
   69: 'Reserva', class Reserva, trigger "DB_OP.DEF05" bit 12
   12: 'Falla térmica en motor Ajuste de ancho de Perfiladores: Comprobar estado de Guardamotor QM07 / DF_QM07 : PROFILEUSE : Moteur OK Axe', class Fallos Perfiladores, trigger "DB_OP.DEF01" bit 3
   6: 'Falla en Control Unit Perfiladores: Comprobar el estado de U13A.3 en el Tablero T02 / DF_VAR04 PROFILEUSE', class Fallos Perfiladores, trigger "DB_OP.DEF01" bit 13
   37: 'Falla al activar alineacion Y de Pieza en Plegadora: Comprobar Sensores 23S5, 23S6, 36S3 y 36S4 + Relé 46K6 / PLIEUSE : DEF MOUVEMENT TAQUAGE Y 46K6 : vérifier 23S5 23S6 36S3 36S4', class Fallos Plegadora, trigger "DB_OP.DEF03" bit 12
   46: 'Falla al Bajar cepillos en Plegadora: Comprobar Sensores 30S7, 30S8, 36S5 y S6S6 + Relé 46K7 / PLIEUSE : DEF MOUVEMENT BROSSE 46K7 : vérifier 30S7 30S8 36S5 S6S6', class Fallos Plegadora, trigger "DB_OP.DEF03" bit 5
   48: 'Reserva', class Reserva, trigger "DB_OP.DEF03" bit 7